// TIA Portal project "GzyHzy_1500" (V15) (continued)
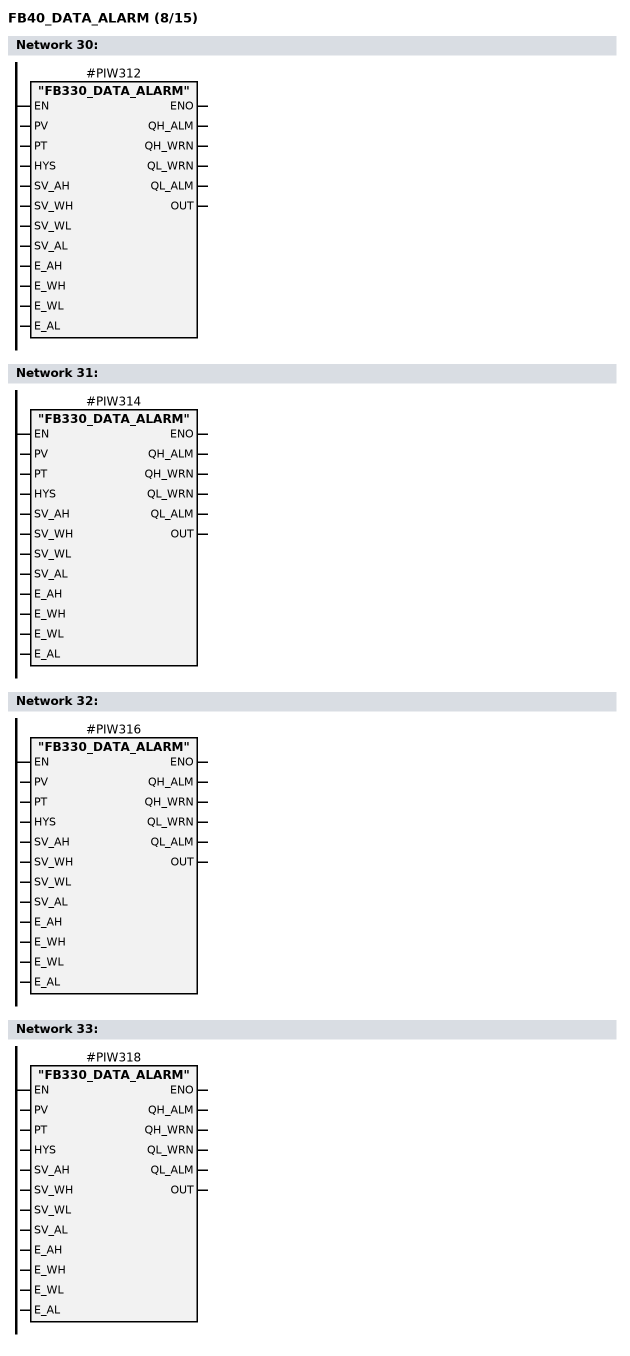
   RUNG wire#powerrail
      #PIW312(PV :=, PT :=, HYS :=, SV_AH :=, SV_WH :=, SV_WL :=, SV_AL :=, E_AH :=, E_WH :=, E_WL :=, E_AL :=, QH_ALM =>, QH_WRN =>, QL_WRN =>, QL_ALM =>, OUT =>)
   END_RUNG
   // the same network as SCL:
   #PIW312();   // "FB330_DATA_ALARM"
END_REGION

REGION Network 31
   RUNG wire#powerrail
      #PIW314(PV :=, PT :=, HYS :=, SV_AH :=, SV_WH :=, SV_WL :=, SV_AL :=, E_AH :=, E_WH :=, E_WL :=, E_AL :=, QH_ALM =>, QH_WRN =>, QL_WRN =>, QL_ALM =>, OUT =>)
   END_RUNG
   // the same network as SCL:
   #PIW314();   // "FB330_DATA_ALARM"
END_REGION

REGION Network 32
   RUNG wire#powerrail
      #PIW316(PV :=, PT :=, HYS :=, SV_AH :=, SV_WH :=, SV_WL :=, SV_AL :=, E_AH :=, E_WH :=, E_WL :=, E_AL :=, QH_ALM =>, QH_WRN =>, QL_WRN =>, QL_ALM =>, OUT =>)
   END_RUNG
   // the same network as SCL:
   #PIW316();   // "FB330_DATA_ALARM"
END_REGION

REGION Network 33
   RUNG wire#powerrail
      #PIW318(PV :=, PT :=, HYS :=, SV_AH :=, SV_WH :=, SV_WL :=, SV_AL :=, E_AH :=, E_WH :=, E_WL :=, E_AL :=, QH_ALM =>, QH_WRN =>, QL_WRN =>, QL_ALM =>, OUT =>)
   END_RUNG
   // the same network as SCL:
   #PIW318();   // "FB330_DATA_ALARM"
END_REGION

REGION Network 34
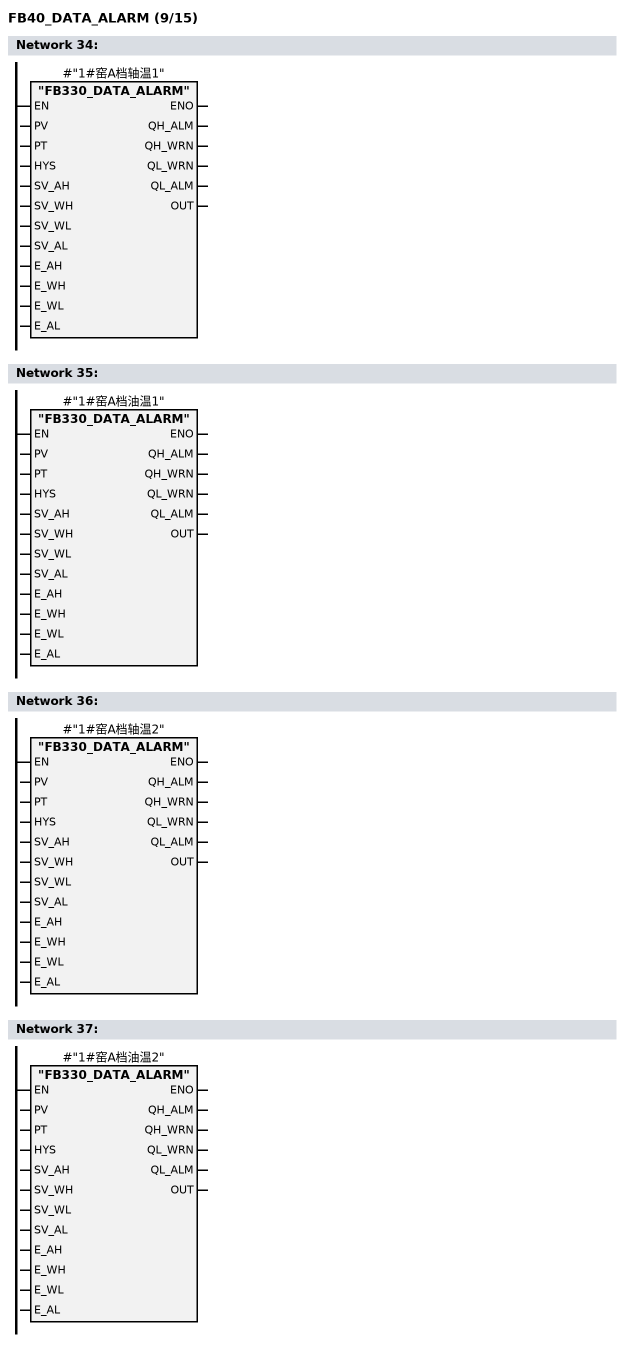
   RUNG wire#powerrail
      #"1#窑A档轴温1"(PV :=, PT :=, HYS :=, SV_AH :=, SV_WH :=, SV_WL :=, SV_AL :=, E_AH :=, E_WH :=, E_WL :=, E_AL :=, QH_ALM =>, QH_WRN =>, QL_WRN =>, QL_ALM =>, OUT =>)
   END_RUNG
   // the same network as SCL:
   #"1#窑A档轴温1"();   // "FB330_DATA_ALARM"
END_REGION

REGION Network 35
   RUNG wire#powerrail
      #"1#窑A档油温1"(PV :=, PT :=, HYS :=, SV_AH :=, SV_WH :=, SV_WL :=, SV_AL :=, E_AH :=, E_WH :=, E_WL :=, E_AL :=, QH_ALM =>, QH_WRN =>, QL_WRN =>, QL_ALM =>, OUT =>)
   END_RUNG
   // the same network as SCL:
   #"1#窑A档油温1"();   // "FB330_DATA_ALARM"
END_REGION

REGION Network 36
   RUNG wire#powerrail
      #"1#窑A档轴温2"(PV :=, PT :=, HYS :=, SV_AH :=, SV_WH :=, SV_WL :=, SV_AL :=, E_AH :=, E_WH :=, E_WL :=, E_AL :=, QH_ALM =>, QH_WRN =>, QL_WRN =>, QL_ALM =>, OUT =>)
   END_RUNG
   // the same network as SCL:
   #"1#窑A档轴温2"();   // "FB330_DATA_ALARM"
END_REGION

REGION Network 37
   RUNG wire#powerrail
      #"1#窑A档油温2"(PV :=, PT :=, HYS :=, SV_AH :=, SV_WH :=, SV_WL :=, SV_AL :=, E_AH :=, E_WH :=, E_WL :=, E_AL :=, QH_ALM =>, QH_WRN =>, QL_WRN =>, QL_ALM =>, OUT =>)
   END_RUNG
   // the same network as SCL:
   #"1#窑A档油温2"();   // "FB330_DATA_ALARM"
END_REGION

REGION Network 38
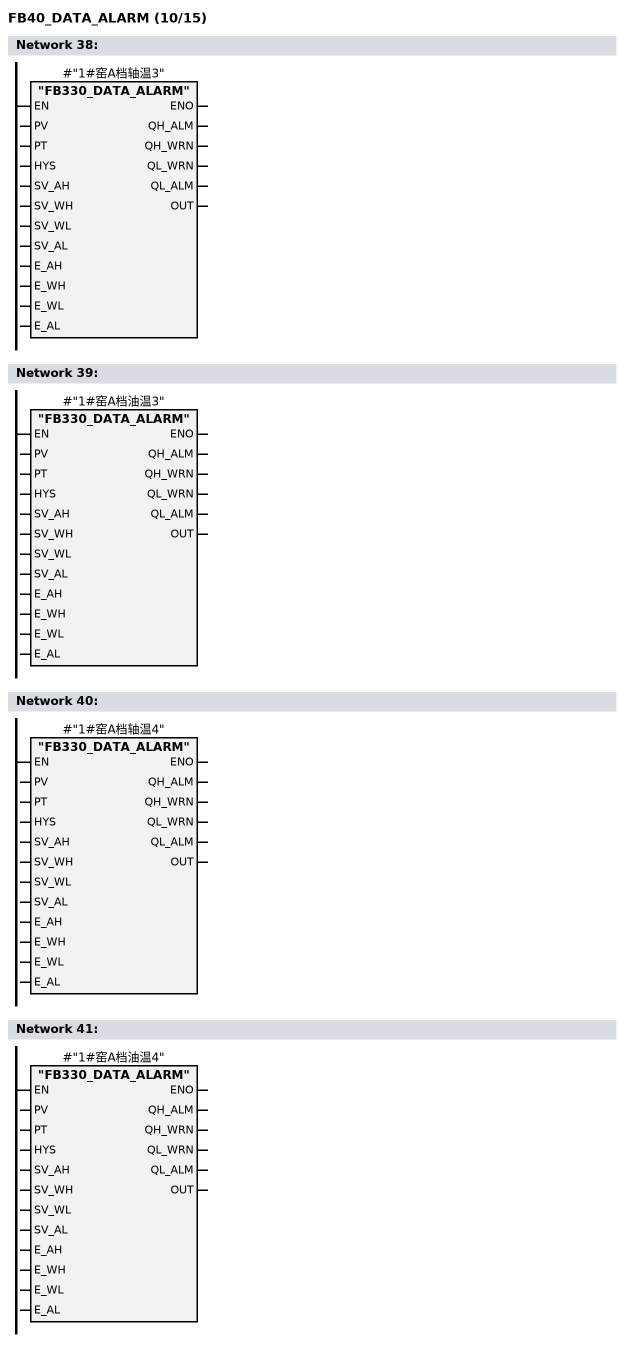
   RUNG wire#powerrail
      #"1#窑A档轴温3"(PV :=, PT :=, HYS :=, SV_AH :=, SV_WH :=, SV_WL :=, SV_AL :=, E_AH :=, E_WH :=, E_WL :=, E_AL :=, QH_ALM =>, QH_WRN =>, QL_WRN =>, QL_ALM =>, OUT =>)
   END_RUNG
   // the same network as SCL:
   #"1#窑A档轴温3"();   // "FB330_DATA_ALARM"
END_REGION

REGION Network 39
   RUNG wire#powerrail
      #"1#窑A档油温3"(PV :=, PT :=, HYS :=, SV_AH :=, SV_WH :=, SV_WL :=, SV_AL :=, E_AH :=, E_WH :=, E_WL :=, E_AL :=, QH_ALM =>, QH_WRN =>, QL_WRN =>, QL_ALM =>, OUT =>)
   END_RUNG
   // the same network as SCL:
   #"1#窑A档油温3"();   // "FB330_DATA_ALARM"
END_REGION

REGION Network 40
   RUNG wire#powerrail
      #"1#窑A档轴温4"(PV :=, PT :=, HYS :=, SV_AH :=, SV_WH :=, SV_WL :=, SV_AL :=, E_AH :=, E_WH :=, E_WL :=, E_AL :=, QH_ALM =>, QH_WRN =>, QL_WRN =>, QL_ALM =>, OUT =>)
   END_RUNG
   // the same network as SCL:
   #"1#窑A档轴温4"();   // "FB330_DATA_ALARM"
END_REGION

REGION Network 41
   RUNG wire#powerrail
      #"1#窑A档油温4"(PV :=, PT :=, HYS :=, SV_AH :=, SV_WH :=, SV_WL :=, SV_AL :=, E_AH :=, E_WH :=, E_WL :=, E_AL :=, QH_ALM =>, QH_WRN =>, QL_WRN =>, QL_ALM =>, OUT =>)
   END_RUNG
   // the same network as SCL:
   #"1#窑A档油温4"();   // "FB330_DATA_ALARM"
END_REGION

REGION Network 42
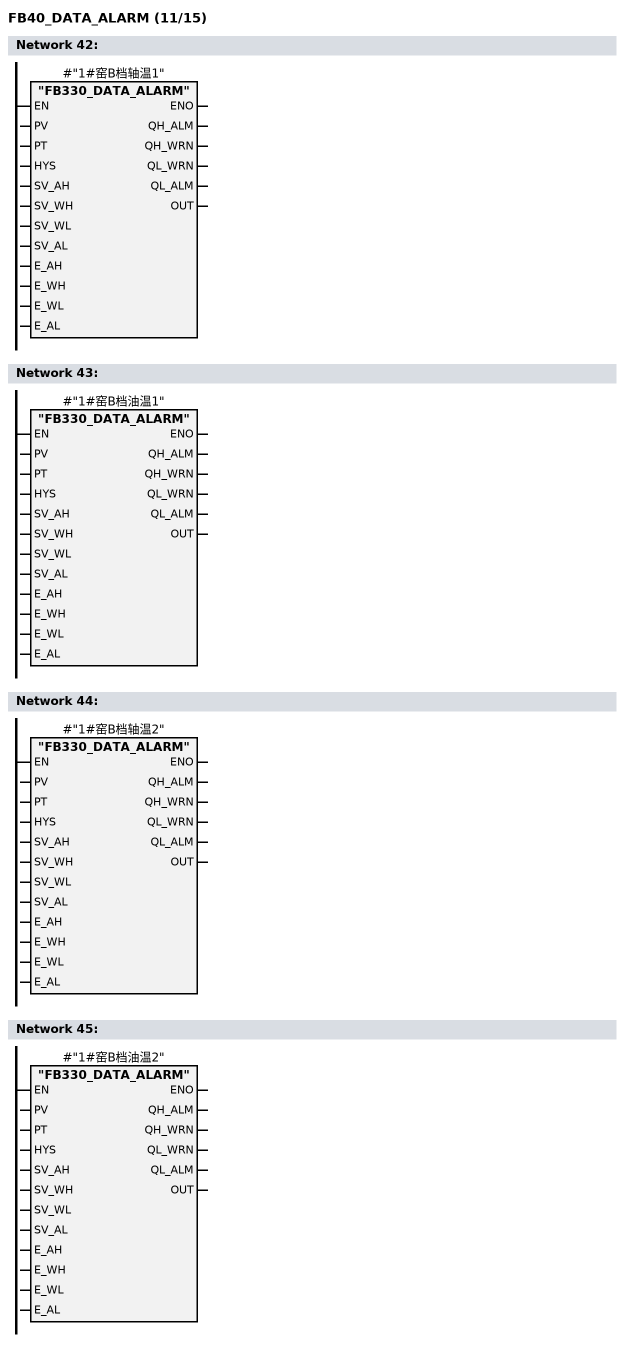
   RUNG wire#powerrail
      #"1#窑B档轴温1"(PV :=, PT :=, HYS :=, SV_AH :=, SV_WH :=, SV_WL :=, SV_AL :=, E_AH :=, E_WH :=, E_WL :=, E_AL :=, QH_ALM =>, QH_WRN =>, QL_WRN =>, QL_ALM =>, OUT =>)
   END_RUNG
   // the same network as SCL:
   #"1#窑B档轴温1"();   // "FB330_DATA_ALARM"
END_REGION

REGION Network 43
   RUNG wire#powerrail
      #"1#窑B档油温1"(PV :=, PT :=, HYS :=, SV_AH :=, SV_WH :=, SV_WL :=, SV_AL :=, E_AH :=, E_WH :=, E_WL :=, E_AL :=, QH_ALM =>, QH_WRN =>, QL_WRN =>, QL_ALM =>, OUT =>)
   END_RUNG
   // the same network as SCL:
   #"1#窑B档油温1"();   // "FB330_DATA_ALARM"
END_REGION

REGION Network 44
   RUNG wire#powerrail
      #"1#窑B档轴温2"(PV :=, PT :=, HYS :=, SV_AH :=, SV_WH :=, SV_WL :=, SV_AL :=, E_AH :=, E_WH :=, E_WL :=, E_AL :=, QH_ALM =>, QH_WRN =>, QL_WRN =>, QL_ALM =>, OUT =>)
   END_RUNG
   // the same network as SCL:
   #"1#窑B档轴温2"();   // "FB330_DATA_ALARM"
END_REGION

REGION Network 45
   RUNG wire#powerrail
      #"1#窑B档油温2"(PV :=, PT :=, HYS :=, SV_AH :=, SV_WH :=, SV_WL :=, SV_AL :=, E_AH :=, E_WH :=, E_WL :=, E_AL :=, QH_ALM =>, QH_WRN =>, QL_WRN =>, QL_ALM =>, OUT =>)
   END_RUNG
   // the same network as SCL:
   #"1#窑B档油温2"();   // "FB330_DATA_ALARM"
END_REGION

REGION Network 46
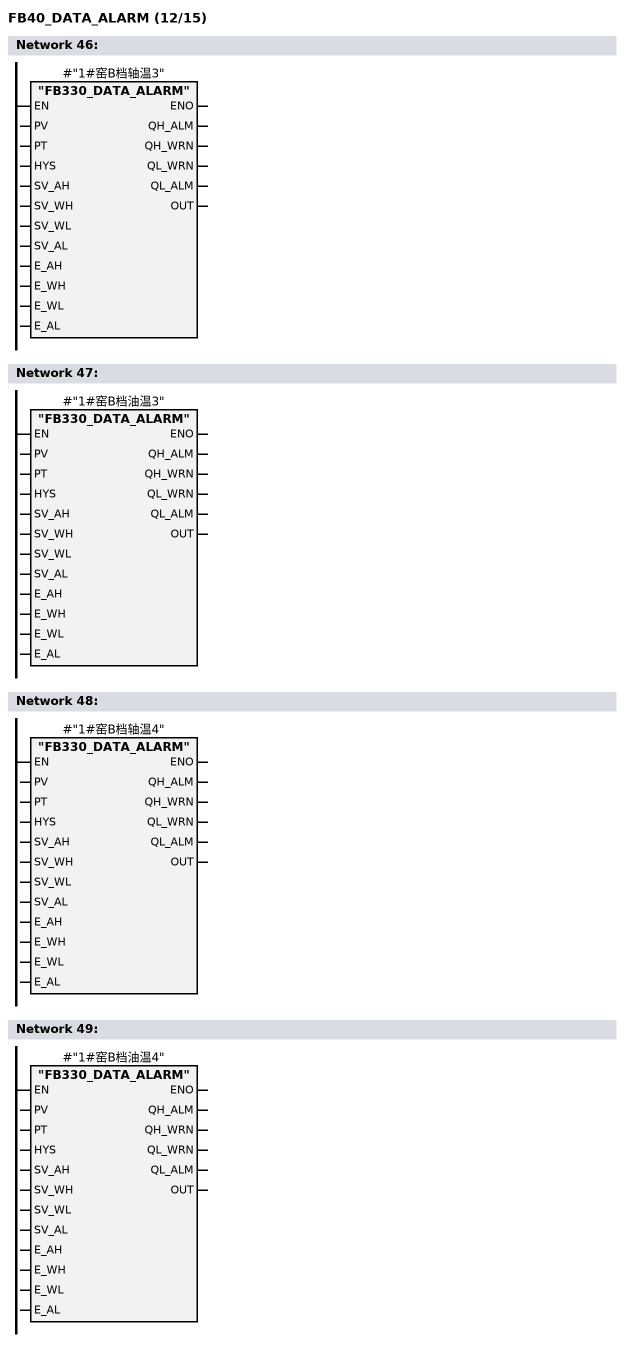
   RUNG wire#powerrail
      #"1#窑B档轴温3"(PV :=, PT :=, HYS :=, SV_AH :=, SV_WH :=, SV_WL :=, SV_AL :=, E_AH :=, E_WH :=, E_WL :=, E_AL :=, QH_ALM =>, QH_WRN =>, QL_WRN =>, QL_ALM =>, OUT =>)
   END_RUNG
   // the same network as SCL:
   #"1#窑B档轴温3"();   // "FB330_DATA_ALARM"
END_REGION

REGION Network 47
   RUNG wire#powerrail
      #"1#窑B档油温3"(PV :=, PT :=, HYS :=, SV_AH :=, SV_WH :=, SV_WL :=, SV_AL :=, E_AH :=, E_WH :=, E_WL :=, E_AL :=, QH_ALM =>, QH_WRN =>, QL_WRN =>, QL_ALM =>, OUT =>)
   END_RUNG
   // the same network as SCL:
   #"1#窑B档油温3"();   // "FB330_DATA_ALARM"
END_REGION

REGION Network 48
   RUNG wire#powerrail
      #"1#窑B档轴温4"(PV :=, PT :=, HYS :=, SV_AH :=, SV_WH :=, SV_WL :=, SV_AL :=, E_AH :=, E_WH :=, E_WL :=, E_AL :=, QH_ALM =>, QH_WRN =>, QL_WRN =>, QL_ALM =>, OUT =>)
   END_RUNG
   // the same network as SCL:
   #"1#窑B档轴温4"();   // "FB330_DATA_ALARM"
END_REGION

REGION Network 49
   RUNG wire#powerrail
      #"1#窑B档油温4"(PV :=, PT :=, HYS :=, SV_AH :=, SV_WH :=, SV_WL :=, SV_AL :=, E_AH :=, E_WH :=, E_WL :=, E_AL :=, QH_ALM =>, QH_WRN =>, QL_WRN =>, QL_ALM =>, OUT =>)
   END_RUNG
   // the same network as SCL:
   #"1#窑B档油温4"();   // "FB330_DATA_ALARM"
END_REGION

REGION Network 50
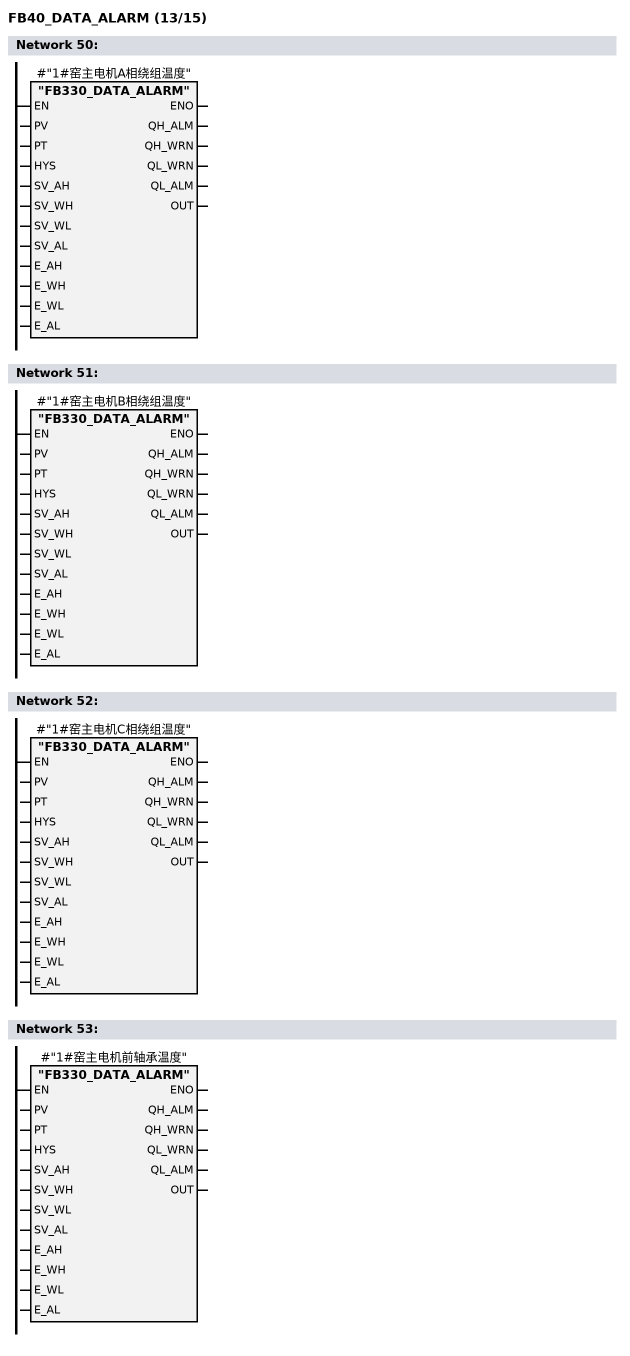
   RUNG wire#powerrail
      #"1#窑主电机A相绕组温度"(PV :=, PT :=, HYS :=, SV_AH :=, SV_WH :=, SV_WL :=, SV_AL :=, E_AH :=, E_WH :=, E_WL :=, E_AL :=, QH_ALM =>, QH_WRN =>, QL_WRN =>, QL_ALM =>, OUT =>)
   END_RUNG
   // the same network as SCL:
   #"1#窑主电机A相绕组温度"();   // "FB330_DATA_ALARM"
END_REGION

REGION Network 51
   RUNG wire#powerrail
      #"1#窑主电机B相绕组温度"(PV :=, PT :=, HYS :=, SV_AH :=, SV_WH :=, SV_WL :=, SV_AL :=, E_AH :=, E_WH :=, E_WL :=, E_AL :=, QH_ALM =>, QH_WRN =>, QL_WRN =>, QL_ALM =>, OUT =>)
   END_RUNG
   // the same network as SCL:
   #"1#窑主电机B相绕组温度"();   // "FB330_DATA_ALARM"
END_REGION

REGION Network 52
   RUNG wire#powerrail
      #"1#窑主电机C相绕组温度"(PV :=, PT :=, HYS :=, SV_AH :=, SV_WH :=, SV_WL :=, SV_AL :=, E_AH :=, E_WH :=, E_WL :=, E_AL :=, QH_ALM =>, QH_WRN =>, QL_WRN =>, QL_ALM =>, OUT =>)
   END_RUNG
   // the same network as SCL:
   #"1#窑主电机C相绕组温度"();   // "FB330_DATA_ALARM"
END_REGION

REGION Network 53
   RUNG wire#powerrail
      #"1#窑主电机前轴承温度"(PV :=, PT :=, HYS :=, SV_AH :=, SV_WH :=, SV_WL :=, SV_AL :=, E_AH :=, E_WH :=, E_WL :=, E_AL :=, QH_ALM =>, QH_WRN =>, QL_WRN =>, QL_ALM =>, OUT =>)
   END_RUNG
   // the same network as SCL:
   #"1#窑主电机前轴承温度"();   // "FB330_DATA_ALARM"
END_REGION

REGION Network 54
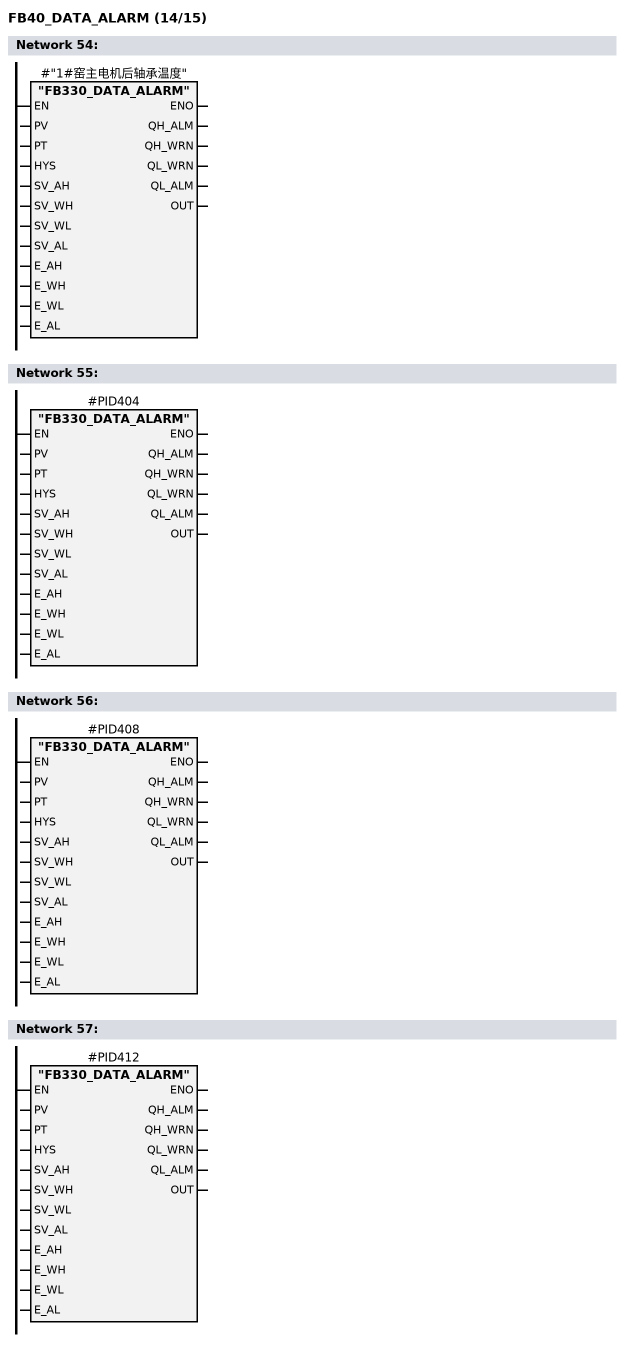
   RUNG wire#powerrail
      #"1#窑主电机后轴承温度"(PV :=, PT :=, HYS :=, SV_AH :=, SV_WH :=, SV_WL :=, SV_AL :=, E_AH :=, E_WH :=, E_WL :=, E_AL :=, QH_ALM =>, QH_WRN =>, QL_WRN =>, QL_ALM =>, OUT =>)
   END_RUNG
   // the same network as SCL:
   #"1#窑主电机后轴承温度"();   // "FB330_DATA_ALARM"
END_REGION

REGION Network 55
   RUNG wire#powerrail
      #PID404(PV :=, PT :=, HYS :=, SV_AH :=, SV_WH :=, SV_WL :=, SV_AL :=, E_AH :=, E_WH :=, E_WL :=, E_AL :=, QH_ALM =>, QH_WRN =>, QL_WRN =>, QL_ALM =>, OUT =>)
   END_RUNG
   // the same network as SCL:
   #PID404();   // "FB330_DATA_ALARM"
END_REGION

REGION Network 56
   RUNG wire#powerrail
      #PID408(PV :=, PT :=, HYS :=, SV_AH :=, SV_WH :=, SV_WL :=, SV_AL :=, E_AH :=, E_WH :=, E_WL :=, E_AL :=, QH_ALM =>, QH_WRN =>, QL_WRN =>, QL_ALM =>, OUT =>)
   END_RUNG
   // the same network as SCL:
   #PID408();   // "FB330_DATA_ALARM"
END_REGION

REGION Network 57
   RUNG wire#powerrail
      #PID412(PV :=, PT :=, HYS :=, SV_AH :=, SV_WH :=, SV_WL :=, SV_AL :=, E_AH :=, E_WH :=, E_WL :=, E_AL :=, QH_ALM =>, QH_WRN =>, QL_WRN =>, QL_ALM =>, OUT =>)
   END_RUNG
   // the same network as SCL:
   #PID412();   // "FB330_DATA_ALARM"
END_REGION

REGION Network 58
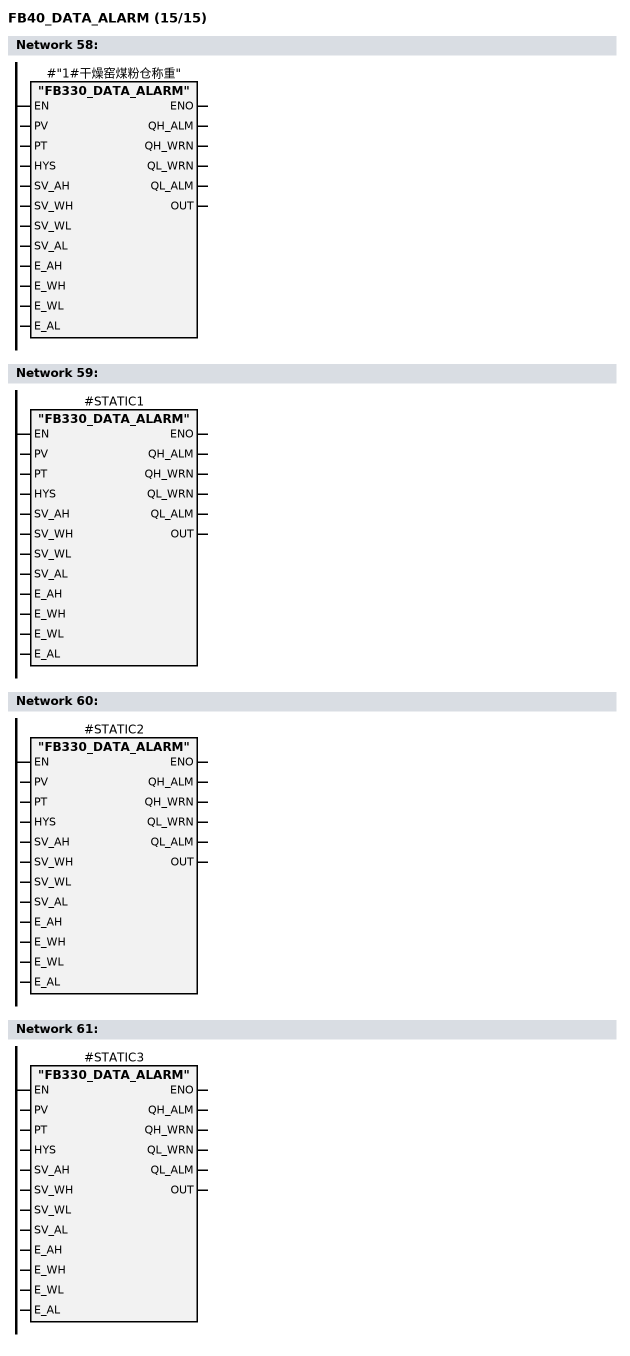
   RUNG wire#powerrail
      #"1#干燥窑煤粉仓称重"(PV :=, PT :=, HYS :=, SV_AH :=, SV_WH :=, SV_WL :=, SV_AL :=, E_AH :=, E_WH :=, E_WL :=, E_AL :=, QH_ALM =>, QH_WRN =>, QL_WRN =>, QL_ALM =>, OUT =>)
   END_RUNG
   // the same network as SCL:
   #"1#干燥窑煤粉仓称重"();   // "FB330_DATA_ALARM"
END_REGION

REGION Network 59
   RUNG wire#powerrail
      #STATIC1(PV :=, PT :=, HYS :=, SV_AH :=, SV_WH :=, SV_WL :=, SV_AL :=, E_AH :=, E_WH :=, E_WL :=, E_AL :=, QH_ALM =>, QH_WRN =>, QL_WRN =>, QL_ALM =>, OUT =>)
   END_RUNG
   // the same network as SCL:
   #STATIC1();   // "FB330_DATA_ALARM"
END_REGION

REGION Network 60
   RUNG wire#powerrail
      #STATIC2(PV :=, PT :=, HYS :=, SV_AH :=, SV_WH :=, SV_WL :=, SV_AL :=, E_AH :=, E_WH :=, E_WL :=, E_AL :=, QH_ALM =>, QH_WRN =>, QL_WRN =>, QL_ALM =>, OUT =>)
   END_RUNG
   // the same network as SCL:
   #STATIC2();   // "FB330_DATA_ALARM"
END_REGION

REGION Network 61
   RUNG wire#powerrail
      #STATIC3(PV :=, PT :=, HYS :=, SV_AH :=, SV_WH :=, SV_WL :=, SV_AL :=, E_AH :=, E_WH :=, E_WL :=, E_AL :=, QH_ALM =>, QH_WRN =>, QL_WRN =>, QL_ALM =>, OUT =>)
   END_RUNG
   // the same network as SCL:
   #STATIC3();   // "FB330_DATA_ALARM"
END_REGION
END_FUNCTION_BLOCK

FUNCTION_BLOCK "FB330_DATA_ALARM"   // FB330, LAD
{ S7_Optimized_Access := 'FALSE' }
VERSION : 0.1
// REAL的报警块
   VAR_INPUT
      PV : Real;   // 过程值
      PT : Real := 1.0;   // 系数
      HYS : Real;   // 回差值
      SV_AH : Real;   // 高报警设定值
      SV_WH : Real;   // 高警告设定值
      SV_WL : Real;   // 低警告设定值
      SV_AL : Real;   // 低报警设定值
      E_AH : Bool;   // 高报警使能
      E_WH : Bool;   // 高警告使能
      E_WL : Bool;   // 低警告使能
      E_AL : Bool;   // 低报警使能
   END_VAR
   VAR_OUTPUT
      QH_ALM : Bool;   // 高报警输出
      QH_WRN : Bool;   // 高警告输出
      QL_WRN : Bool;   // 低警告输出
      QL_ALM : Bool;   // 低报警输出
      OUT : Real;   // 输出
   END_VAR
   VAR
      SR1 : Bool;
      SR2 : Bool;
      SR3 : Bool;
      SR4 : Bool;
   END_VAR
   VAR_TEMP
      TEMP_AH : Real;
      TEMP_WH : Real;
      TEMP_AL : Real;
      TEMP_WL : Real;
      TEMP_OUT : Real;
   END_VAR
BEGIN

REGION Network 1
   // 系数转换
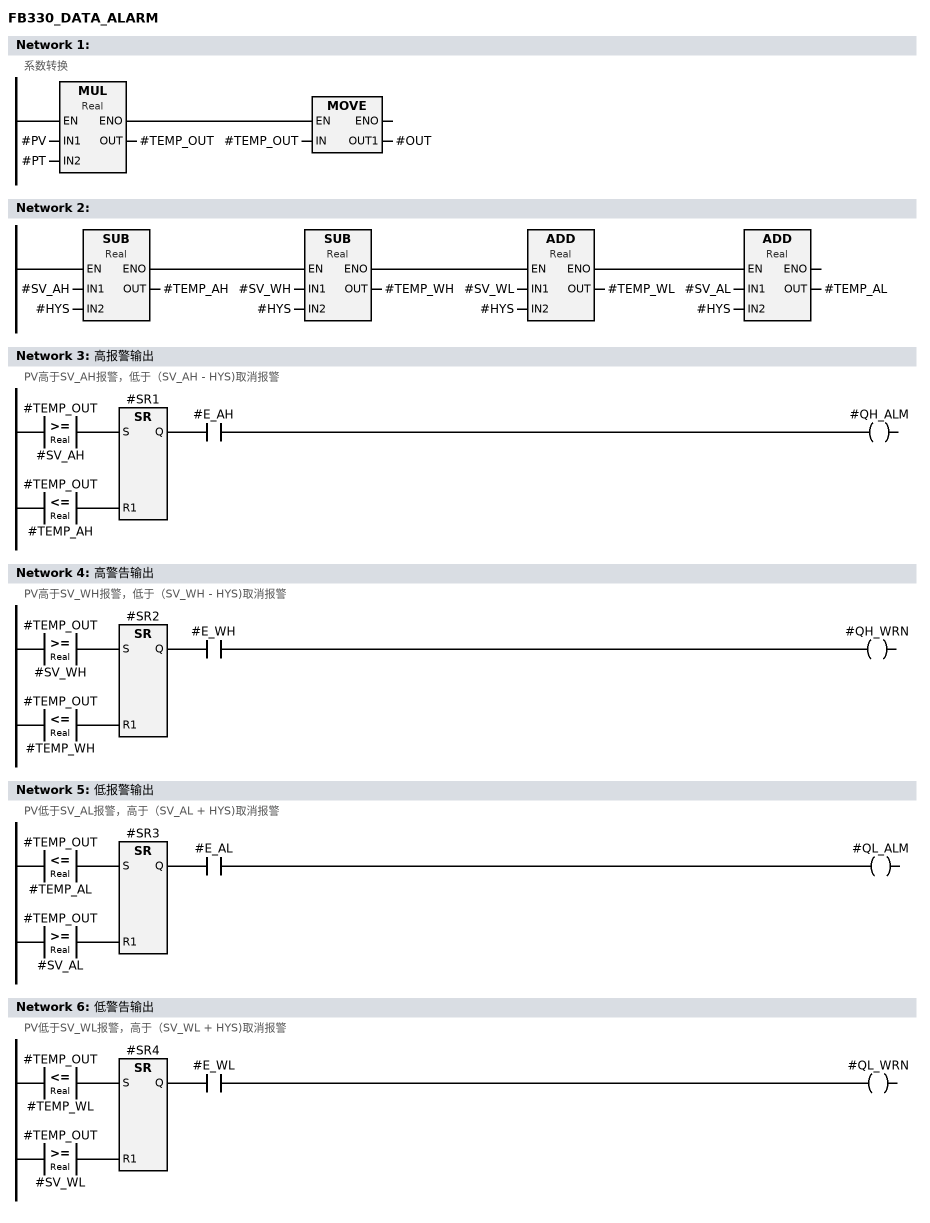
   RUNG wire#powerrail
      { S7_Templates := "SrcType := Real"; S7_GenerateENO := "TRUE" } Mul(in1 := #PV, in2 := #PT, out => #TEMP_OUT)
      { S7_GenerateENO := "TRUE" } Move(in := #TEMP_OUT, out1 => #OUT)
   END_RUNG
   // the same network as SCL:
   // ENO of a box is taken as its EN; it also drops when the box reports an error
   #TEMP_OUT := #PV * #PT;
   #OUT := #TEMP_OUT;
END_REGION

REGION Network 2
   RUNG wire#powerrail
      { S7_Templates := "SrcType := Real"; S7_GenerateENO := "TRUE" } Sub(in1 := #SV_AH, in2 := #HYS, out => #TEMP_AH)
      { S7_Templates := "SrcType := Real"; S7_GenerateENO := "TRUE" } Sub(in1 := #SV_WH, in2 := #HYS, out => #TEMP_WH)
      { S7_Templates := "SrcType := Real"; S7_GenerateENO := "TRUE" } Add(in1 := #SV_WL, in2 := #HYS, out => #TEMP_WL)
      { S7_Templates := "SrcType := Real"; S7_GenerateENO := "TRUE" } Add(in1 := #SV_AL, in2 := #HYS, out => #TEMP_AL)
   END_RUNG
   // the same network as SCL:
   // ENO of a box is taken as its EN; it also drops when the box reports an error
   #TEMP_AH := #SV_AH - #HYS;
   #TEMP_WH := #SV_WH - #HYS;
   #TEMP_WL := #SV_WL + #HYS;
   #TEMP_AL := #SV_AL + #HYS;
END_REGION

REGION Network 3: 高报警输出
   // PV高于SV_AH报警，低于（SV_AH - HYS)取消报警
   RUNG wire#powerrail
      { S7_Templates := "SrcType := Real" } GE_Contact(in1 := #TEMP_OUT, in2 := #SV_AH)
      S_SR(operand := #SR1, r1 := wire#w1)
      Contact( #E_AH )
      Coil( #QH_ALM )
   END_RUNG
   RUNG wire#powerrail
      { S7_Templates := "SrcType := Real" } LE_Contact(in1 := #TEMP_OUT, in2 := #TEMP_AH)
   END_RUNG wire#w1
   // the same network as SCL:
   IF #TEMP_OUT >= #SV_AH THEN
       #SR1 := TRUE;   // SR flip-flop
   END_IF;
   IF #TEMP_OUT <= #TEMP_AH THEN #SR1 := FALSE; END_IF;
   #QH_ALM := #SR1 AND #E_AH;
END_REGION

REGION Network 4: 高警告输出
   // PV高于SV_WH报警，低于（SV_WH - HYS)取消报警
   RUNG wire#powerrail
      { S7_Templates := "SrcType := Real" } GE_Contact(in1 := #TEMP_OUT, in2 := #SV_WH)
      S_SR(operand := #SR2, r1 := wire#w1)
      Contact( #E_WH )
      Coil( #QH_WRN )
   END_RUNG
   RUNG wire#powerrail
      { S7_Templates := "SrcType := Real" } LE_Contact(in1 := #TEMP_OUT, in2 := #TEMP_WH)
   END_RUNG wire#w1
   // the same network as SCL:
   IF #TEMP_OUT >= #SV_WH THEN
       #SR2 := TRUE;   // SR flip-flop
   END_IF;
   IF #TEMP_OUT <= #TEMP_WH THEN #SR2 := FALSE; END_IF;
   #QH_WRN := #SR2 AND #E_WH;
END_REGION

REGION Network 5: 低报警输出
   // PV低于SV_AL报警，高于（SV_AL + HYS)取消报警
   RUNG wire#powerrail
      { S7_Templates := "SrcType := Real" } LE_Contact(in1 := #TEMP_OUT, in2 := #TEMP_AL)
      S_SR(operand := #SR3, r1 := wire#w1)
      Contact( #E_AL )
      Coil( #QL_ALM )
   END_RUNG
   RUNG wire#powerrail
      { S7_Templates := "SrcType := Real" } GE_Contact(in1 := #TEMP_OUT, in2 := #SV_AL)
   END_RUNG wire#w1
   // the same network as SCL:
   IF #TEMP_OUT <= #TEMP_AL THEN
       #SR3 := TRUE;   // SR flip-flop
   END_IF;
   IF #TEMP_OUT >= #SV_AL THEN #SR3 := FALSE; END_IF;
   #QL_ALM := #SR3 AND #E_AL;
END_REGION

REGION Network 6: 低警告输出
   // PV低于SV_WL报警，高于（SV_WL + HYS)取消报警
   RUNG wire#powerrail
      { S7_Templates := "SrcType := Real" } LE_Contact(in1 := #TEMP_OUT, in2 := #TEMP_WL)
      S_SR(operand := #SR4, r1 := wire#w1)
      Contact( #E_WL )
      Coil( #QL_WRN )
   END_RUNG
   RUNG wire#powerrail
      { S7_Templates := "SrcType := Real" } GE_Contact(in1 := #TEMP_OUT, in2 := #SV_WL)
   END_RUNG wire#w1
   // the same network as SCL:
   IF #TEMP_OUT <= #TEMP_WL THEN
       #SR4 := TRUE;   // SR flip-flop
   END_IF;
   IF #TEMP_OUT >= #SV_WL THEN #SR4 := FALSE; END_IF;
   #QL_WRN := #SR4 AND #E_WL;
END_REGION
END_FUNCTION_BLOCK

FUNCTION_BLOCK "累计功能块2"   // FB333, LAD
{ S7_Optimized_Access := 'FALSE' }
VERSION : 0.1
   VAR_INPUT
      PV : Real;
      CLEAR1 : Bool;
      CLEAR2 : Bool;
      CLEAR3 : Bool;
      CLEAR4 : Bool;
   END_VAR
   VAR_OUTPUT
      OUT1 : Real;
      OUT2 : Real;
      OUT3 : Real;
      OUT4 : Real;
   END_VAR
   VAR
      "REAL" : Real;
      REAL1_1 : Real;
      REAL1_2 : Real;
      REAL1_3 : Real;
      REAL2_1 : Real;
      REAL2_2 : Real;
      REAL2_3 : Real;
      REAL3_1 : Real;
      REAL3_2 : Real;
      REAL3_3 : Real;
      REAL4_1 : Real;
      REAL4_2 : Real;
      REAL4_3 : Real;
      PV_DINT : DInt;
      DINT1 : DInt;
      DINT2 : DInt;
      DINT3 : DInt;
      DINT4 : DInt;
      P1 : Bool;
      P2 : Bool;
      P3 : Bool;
      P4 : Bool;
   END_VAR
   VAR_TEMP   // added for the SCL form of the ladder/FBD networks
      _w1 : Bool;
      _w2 : Bool;
   END_VAR
BEGIN

REGION Network 1
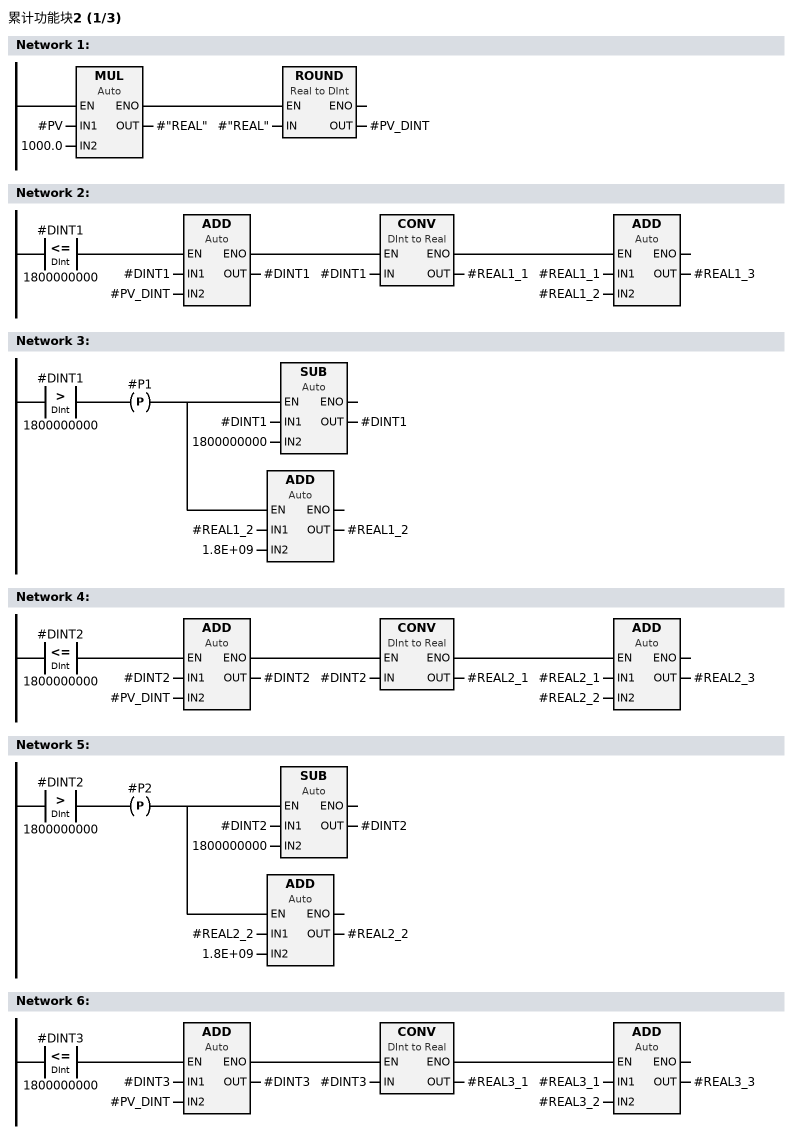
   RUNG wire#powerrail
      Mul(in1 := #PV, in2 := 1000.0, out => #"REAL")
      { S7_Templates := "[SrcType := Real, DestType := DInt]" } Round(in := #"REAL", out => #PV_DINT)
   END_RUNG
   // the same network as SCL:
   #"REAL" := #PV * 1000.0;
   #PV_DINT := ROUND(#"REAL");
END_REGION

REGION Network 2
   RUNG wire#powerrail
      { S7_Templates := "SrcType := DInt" } LE_Contact(in1 := #DINT1, in2 := 1800000000)
      Add(in1 := #DINT1, in2 := #PV_DINT, out => #DINT1)
      { S7_Templates := "[SrcType := DInt, DestType := Real]" } Convert(in := #DINT1, out => #REAL1_1)
      Add(in1 := #REAL1_1, in2 := #REAL1_2, out => #REAL1_3)
   END_RUNG
   // the same network as SCL:
   #_w1 := #DINT1 <= 1800000000;
   IF #_w1 THEN
       #DINT1 := #DINT1 + #PV_DINT;
       #REAL1_1 := DINT_TO_REAL(#DINT1);
       #REAL1_3 := #REAL1_1 + #REAL1_2;
   END_IF;
END_REGION

REGION Network 3
   RUNG wire#powerrail
      { S7_Templates := "SrcType := DInt" } GT_Contact(in1 := #DINT1, in2 := 1800000000)
      P_Trig( #P1 )
      wire#w1
      Sub(in1 := #DINT1, in2 := 1800000000, out => #DINT1)
   END_RUNG
   RUNG wire#w1
      Add(in1 := #REAL1_2, in2 := 1.8E+09, out => #REAL1_2)
   END_RUNG
   // the same network as SCL:
   #_w1 := #DINT1 > 1800000000;
   #_w2 := #_w1 AND NOT #P1;   // rising edge
   #P1 := #_w1;
   IF #_w2 THEN
       #DINT1 := #DINT1 - 1800000000;
       #REAL1_2 := #REAL1_2 + 1.8E+09;
   END_IF;
END_REGION

REGION Network 4
   RUNG wire#powerrail
      { S7_Templates := "SrcType := DInt" } LE_Contact(in1 := #DINT2, in2 := 1800000000)
      Add(in1 := #DINT2, in2 := #PV_DINT, out => #DINT2)
      { S7_Templates := "[SrcType := DInt, DestType := Real]" } Convert(in := #DINT2, out => #REAL2_1)
      Add(in1 := #REAL2_1, in2 := #REAL2_2, out => #REAL2_3)
   END_RUNG
   // the same network as SCL:
   #_w1 := #DINT2 <= 1800000000;
   IF #_w1 THEN
       #DINT2 := #DINT2 + #PV_DINT;
       #REAL2_1 := DINT_TO_REAL(#DINT2);
       #REAL2_3 := #REAL2_1 + #REAL2_2;
   END_IF;
END_REGION

REGION Network 5
   RUNG wire#powerrail
      { S7_Templates := "SrcType := DInt" } GT_Contact(in1 := #DINT2, in2 := 1800000000)
      P_Trig( #P2 )
      wire#w1
      Sub(in1 := #DINT2, in2 := 1800000000, out => #DINT2)
   END_RUNG
   RUNG wire#w1
      Add(in1 := #REAL2_2, in2 := 1.8E+09, out => #REAL2_2)
   END_RUNG
   // the same network as SCL:
   #_w1 := #DINT2 > 1800000000;
   #_w2 := #_w1 AND NOT #P2;   // rising edge
   #P2 := #_w1;
   IF #_w2 THEN
       #DINT2 := #DINT2 - 1800000000;
       #REAL2_2 := #REAL2_2 + 1.8E+09;
   END_IF;
END_REGION

REGION Network 6
   RUNG wire#powerrail
      { S7_Templates := "SrcType := DInt" } LE_Contact(in1 := #DINT3, in2 := 1800000000)
      Add(in1 := #DINT3, in2 := #PV_DINT, out => #DINT3)
      { S7_Templates := "[SrcType := DInt, DestType := Real]" } Convert(in := #DINT3, out => #REAL3_1)
      Add(in1 := #REAL3_1, in2 := #REAL3_2, out => #REAL3_3)
   END_RUNG
   // the same network as SCL:
   #_w1 := #DINT3 <= 1800000000;
   IF #_w1 THEN
       #DINT3 := #DINT3 + #PV_DINT;
       #REAL3_1 := DINT_TO_REAL(#DINT3);
       #REAL3_3 := #REAL3_1 + #REAL3_2;
   END_IF;
END_REGION

REGION Network 7
